(* Logix 5000 project; controller MV vendor 1 type 14 code 217 rev 31.11; software revision 31.00; part 42 of 53 *)
(* tags used below, declared in another part *)
   Always_Off : BOOL;
   Dummy : BOOL;
   MV20_TP_Capture_Volume_Timer : TIMER;
   MV_BM01_AV01_CIP : BOOL;
   MV_data_file_value_to_move : DINT;
   MV_Enable_MV20_NewPressureControl : BOOL;
   MV_from_data_file : DINT;
   MV_from_data_offset : DINT;
   MV_MV10_RTD1_AI : PlantItem;   // MV10_RTD1
   MV_MV11_RTD1_AI : PlantItem;   // MV11_RTD1
   MV_MV12_RTD1_AI : PlantItem;   // MV12_RTD1
   MV_MV13_RTD1_AI : PlantItem;   // MV13_RTD1
   MV_MV14_RTD1_AI : PlantItem;   // MV14_RTD1
   MV_MV15_RTD1_AI : PlantItem;   // MV15_RTD1
   MV_MV16_RTD1_AI : PlantItem;   // MV16_RTD1
   MV_MV17_RTD1_AI : PlantItem;   // MV17_RTD1
   MV_MV18_RTD1_AI : PlantItem;   // MV18_RTD1
   MV_MV19_RTD1_AI : PlantItem;   // MV19_RTD1
   MV_MV1_RTD1_AI : PlantItem;   // MV1_RTD1
   MV_MV20_CO2_ON_PreStorage : BOOL;
   MV_MV20_CO2_ON_Storage : BOOL;
   MV_MV20_Filling_PulseLevel : REAL;
   MV_MV20_LTX07_TrueLevel : REAL;
   MV_MV20_ProxiesOK : BOOL;
   MV_MV20_PTX01_AI : PlantItem;   // MV20_PTX01
   MV_MV20_RTD1_AI : PlantItem;   // MV20_RTD1
   MV_MV20_TP_Command : DINT;
   MV_MV20_TP_Dirty : BOOL;
   MV_MV20_TP_Emptying_Level_Setpoint : REAL;
   MV_MV20_TP_Idle : BOOL;
   MV_MV20_TP_KBDepressure : BOOL;
   MV_MV20_TP_KBFilling : BOOL;
   MV_MV20_TP_KBFilling_M : BOOL;
   MV_MV20_TP_KBPreEmptyPressure : BOOL;
   MV_MV20_TP_KBPrePressurise : BOOL;
   MV_MV20_TP_KBPurgeFromTop : BOOL;
   MV_MV20_TP_KBPurgeTimer : TIMER;
   MV_MV20_TP_KBStorage : BOOL;
   MV_MV20_TP_ONS : BOOL;
   MV_MV20_TP_Prompt : DINT;
   MV_MV20_TP_ReadyToFillKB : BOOL;
   MV_MV20_TP_ReadyToFillKB_M : BOOL;
   MV_MV20_TP_Running : BOOL;
   MV_MV20_TP_Setpoint : REAL;
   MV_MV20_TP_Status : DINT;   // 0 = Idle, 1 = Running, 2 = Held, 3 = Faulted
   MV_MV20_TP_Step : DINT;
   MV_MV20_TP_Steptime : DINT;
   MV_MV20_TP_UpperLimit : REAL;
   MV_MV20_Transfer_StartLevel : REAL;
   MV_MV21_RTD1_AI : PlantItem;   // MV21_RTD1
   MV_MV22_RTD1_AI : PlantItem;   // MV22_RTD1
   MV_MV23_RTD1_AI : PlantItem;   // MV23_RTD1
   MV_MV2_RTD1_AI : PlantItem;   // MV2_RTD1
   MV_MV30_RTD1_AI : PlantItem;   // MV30_RTD1
   MV_MV31_RTD1_AI : PlantItem;   // MV31_RTD1
   MV_MV32_RTD1_AI : PlantItem;   // MV32_RTD1
   MV_MV33_RTD1_AI : PlantItem;   // MV33_RTD1
   MV_MV34_RTD1_AI : PlantItem;   // MV34_RTD1
   MV_MV35_RTD1_AI : PlantItem;   // MV35_RTD1
   MV_MV36_TTX01_AI : PlantItem;   // MV36_TTX01
   MV_MV37_TTX01_AI : PlantItem;   // MV37_TTX01
   MV_MV38_TTX01_AI : PlantItem;   // MV38_TTX01
   MV_MV39_TTX01_AI : PlantItem;   // MV39_TTX01
   MV_MV3_RTD1_AI : PlantItem;   // MV3_RTD1
   MV_MV40_TTX01_AI : PlantItem;   // MV40_TTX01
   MV_MV41_TTX01_AI : PlantItem;   // MV41_TTX01
   MV_MV42_TTX01_AI : PlantItem;   // MV42_TTX01
   MV_MV43_TTX01_AI : PlantItem;   // MV43_TTX01
   MV_MV44_TTX01_AI : PlantItem;   // MV44_TTX01
   MV_MV45_TTX01_AI : PlantItem;   // MV45_TTX01
   MV_MV46_TTX01_AI : PlantItem;   // MV46_TTX01
   MV_MV47_TTX01_AI : PlantItem;   // MV47_TTX01
   MV_MV4_RTD1_AI : PlantItem;   // MV4_RTD1
   MV_MV5_RTD1_AI : PlantItem;   // MV5_RTD1
   MV_MV6_RTD1_AI : PlantItem;   // MV6_RTD1
   MV_MV7_RTD1_AI : PlantItem;   // MV7_RTD1
   MV_MV8_RTD1_AI : PlantItem;   // MV8_RTD1
   MV_MV9_RTD1_AI : PlantItem;   // MV9_RTD1
   MV_N106 : INT[255];   // ROUSE_BUFF Rouser control vesse l data buffer
   MV_N110 : INT[255];   // MV DATA 0 CURRENT FV DATA
   MV_N111 : INT[50];   // MV 1, CURRENT FV DATA
   MV_N112 : INT[50];   // MV 2, CURRENT FV DATA
   MV_N113 : INT[50];   // MV 3, CURRENT FV DATA
   MV_N114 : INT[50];   // MV 4, CURRENT FV DATA
   MV_N115 : INT[50];   // MV 5, CURRENT FV DATA
   MV_N116 : INT[50];   // MV 6, CURRENT FV DATA
   MV_N117 : INT[50];   // MV 7, CURRENT FV DATA
   MV_N118 : INT[50];   // MV 8, CURRENT FV DATA
   MV_N119 : INT[50];   // MV 9, CURRENT FV DATA
   MV_N120 : INT[50];   // MV 10, CURRENT FV DATA
   MV_N121 : INT[50];   // MV 11, CURRENT FV DATA
   MV_N122 : INT[50];   // MV 12, CURRENT FV DATA
   MV_N123 : INT[50];   // MV 13, CURRENT FV DATA
   MV_N124 : INT[50];   // MV 14, CURRENT FV DATA
   MV_N125 : INT[50];   // MV 15, CURRENT FV DATA
   MV_N126 : INT[50];   // MV 16, CURRENT FV DATA
   MV_N127 : INT[50];   // MV 17, CURRENT FV DATA
   MV_N128 : INT[50];   // MV 18, CURRENT FV DATA
   MV_N129 : INT[50];   // MV 19, CURRENT FV DATA
   MV_N130 : INT[50];   // MV 30, CURRENT FV DATA
   MV_N131 : INT[50];   // MV 31, CURRENT FV DATA
   MV_N132 : INT[50];   // MV 32, CURRENT FV DATA
   MV_N133 : INT[50];   // MV 33, CURRENT FV DATA
   MV_N134 : INT[50];   // MV 34, CURRENT FV DATA
   MV_N135 : INT[50];   // MV 35, CURRENT FV DATA
   MV_N136 : INT[50];   // MV 20, CURRENT FV DATA
   MV_N137 : INT[50];   // MV 21, CURRENT FV DATA
   MV_N138 : INT[50];   // MV 22, CURRENT FV DATA
   MV_N139 : INT[50];   // MV 23, CURRENT FV DATA
   MV_N140 : INT[50];   // MV 36, CURRENT FV DATA
   MV_N141 : INT[50];   // MV 37, CURRENT FV DATA
   MV_N142 : INT[50];   // MV 38, CURRENT FV DATA
   MV_N143 : INT[50];   // MV 39, CURRENT FV DATA
   MV_N144 : INT[50];   // MV 40, CURRENT FV DATA
   MV_N145 : INT[50];   // MV 41, CURRENT FV DATA
   MV_N146 : INT[50];   // MV 42, CURRENT FV DATA
   MV_N147 : INT[50];   // MV 43, CURRENT FV DATA
   MV_N148 : INT[50];   // MV 44, CURRENT FV DATA
   MV_N149 : INT[50];   // MV 45, CURRENT FV DATA
   MV_N150 : INT[50];   // MV 36, CURRENT FV DATA
   MV_N151 : INT[50];   // MV 47, CURRENT FV DATA
   MV_TP_CaskPrefillPressure : REAL;
   MV_TP_Emptying_Volume_Setpoint : REAL;
   MV_TP_KBEmptyingPressure : REAL;
   MV_TP_KBFillingPressure : REAL;
   MV_TP_KBPrefillPressure : REAL;
   MV_TP_KBStoragePressure : REAL;
   MV_TP_KBStoragePressureLevel : REAL;
   MV_TP_NoCIPDelay : DINT;
(* MV_Common, continued *)

ROUTINE MV_Get_FV_Datafile_Value   (* ladder *)
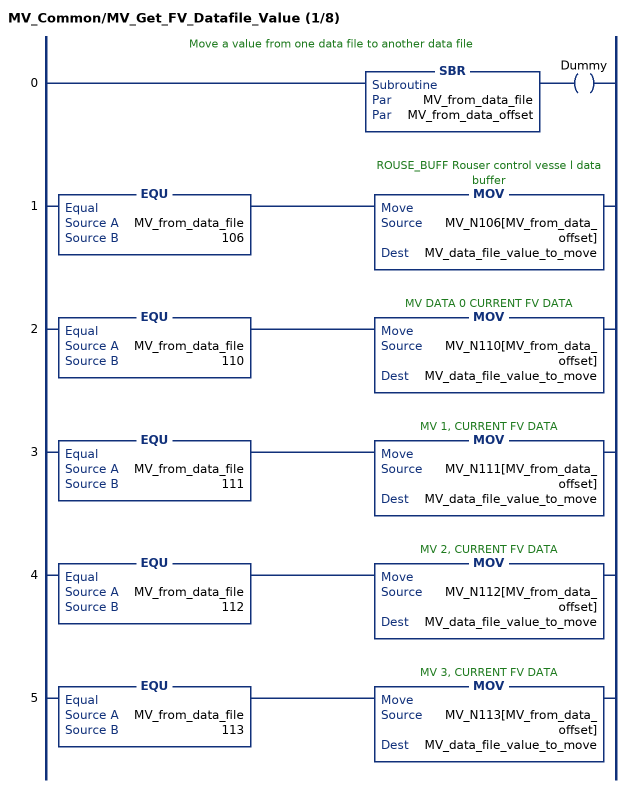
   // Move a value from one data file to another data file
   0: SBR(MV_from_data_file,MV_from_data_offset)OTE(Dummy);
   1: EQU(MV_from_data_file,106)MOV(MV_N106[MV_from_data_offset],MV_data_file_value_to_move);
   2: EQU(MV_from_data_file,110)MOV(MV_N110[MV_from_data_offset],MV_data_file_value_to_move);
   3: EQU(MV_from_data_file,111)MOV(MV_N111[MV_from_data_offset],MV_data_file_value_to_move);
   4: EQU(MV_from_data_file,112)MOV(MV_N112[MV_from_data_offset],MV_data_file_value_to_move);
   5: EQU(MV_from_data_file,113)MOV(MV_N113[MV_from_data_offset],MV_data_file_value_to_move);
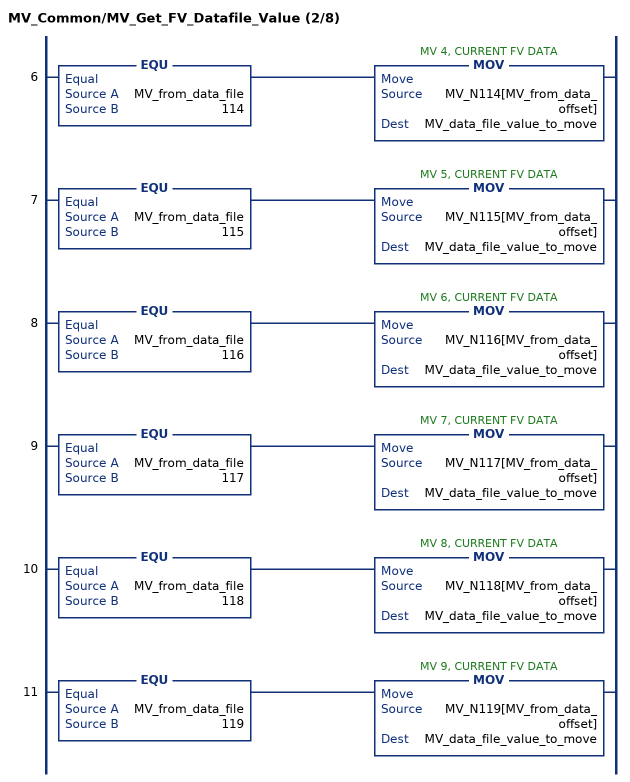
   6: EQU(MV_from_data_file,114)MOV(MV_N114[MV_from_data_offset],MV_data_file_value_to_move);
   7: EQU(MV_from_data_file,115)MOV(MV_N115[MV_from_data_offset],MV_data_file_value_to_move);
   8: EQU(MV_from_data_file,116)MOV(MV_N116[MV_from_data_offset],MV_data_file_value_to_move);
   9: EQU(MV_from_data_file,117)MOV(MV_N117[MV_from_data_offset],MV_data_file_value_to_move);
   10: EQU(MV_from_data_file,118)MOV(MV_N118[MV_from_data_offset],MV_data_file_value_to_move);
   11: EQU(MV_from_data_file,119)MOV(MV_N119[MV_from_data_offset],MV_data_file_value_to_move);
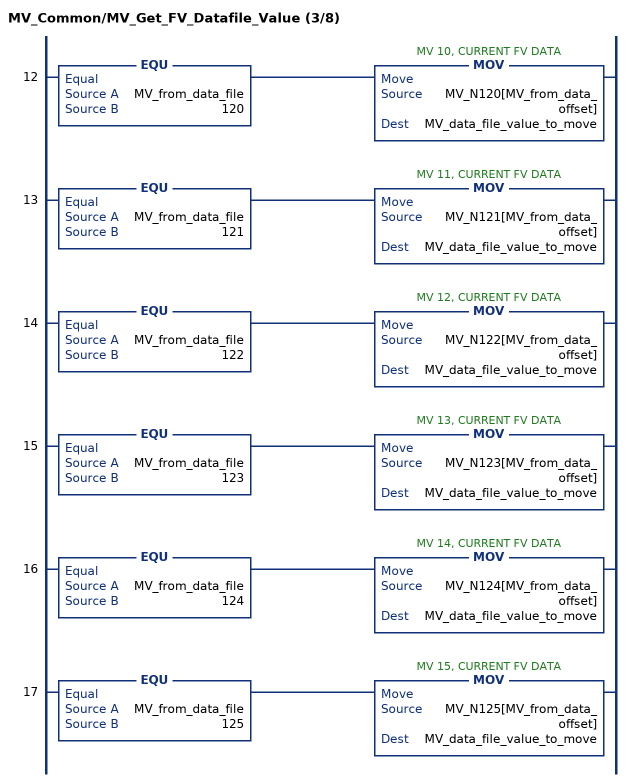
   12: EQU(MV_from_data_file,120)MOV(MV_N120[MV_from_data_offset],MV_data_file_value_to_move);
   13: EQU(MV_from_data_file,121)MOV(MV_N121[MV_from_data_offset],MV_data_file_value_to_move);
   14: EQU(MV_from_data_file,122)MOV(MV_N122[MV_from_data_offset],MV_data_file_value_to_move);
   15: EQU(MV_from_data_file,123)MOV(MV_N123[MV_from_data_offset],MV_data_file_value_to_move);
   16: EQU(MV_from_data_file,124)MOV(MV_N124[MV_from_data_offset],MV_data_file_value_to_move);
   17: EQU(MV_from_data_file,125)MOV(MV_N125[MV_from_data_offset],MV_data_file_value_to_move);
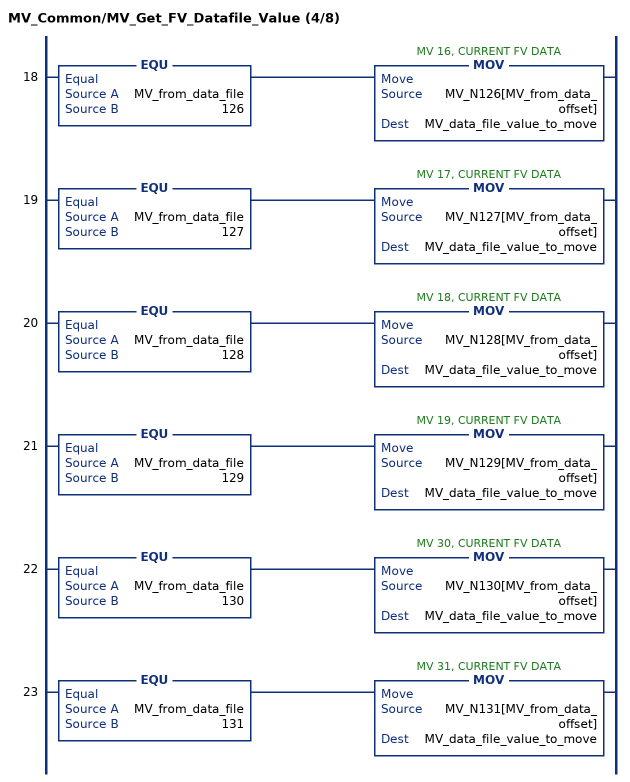
   18: EQU(MV_from_data_file,126)MOV(MV_N126[MV_from_data_offset],MV_data_file_value_to_move);
   19: EQU(MV_from_data_file,127)MOV(MV_N127[MV_from_data_offset],MV_data_file_value_to_move);
   20: EQU(MV_from_data_file,128)MOV(MV_N128[MV_from_data_offset],MV_data_file_value_to_move);
   21: EQU(MV_from_data_file,129)MOV(MV_N129[MV_from_data_offset],MV_data_file_value_to_move);
   22: EQU(MV_from_data_file,130)MOV(MV_N130[MV_from_data_offset],MV_data_file_value_to_move);
   23: EQU(MV_from_data_file,131)MOV(MV_N131[MV_from_data_offset],MV_data_file_value_to_move);
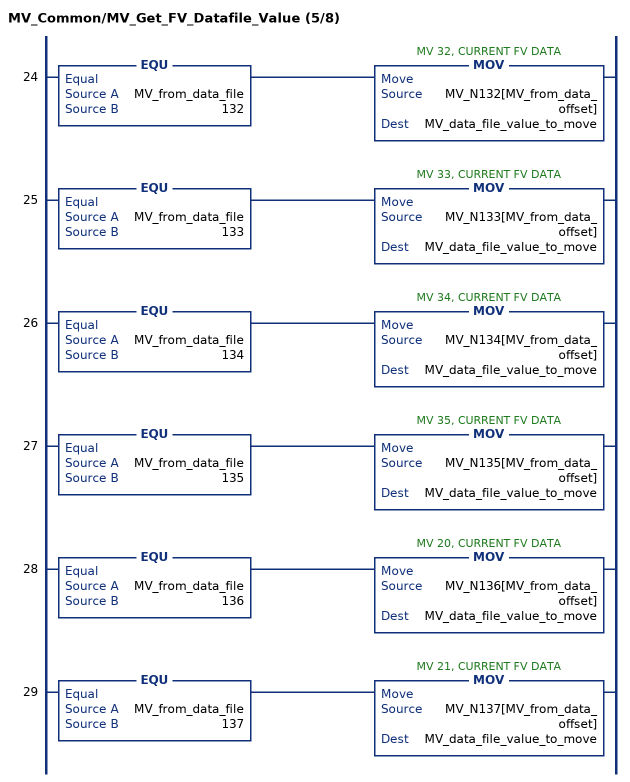
   24: EQU(MV_from_data_file,132)MOV(MV_N132[MV_from_data_offset],MV_data_file_value_to_move);
   25: EQU(MV_from_data_file,133)MOV(MV_N133[MV_from_data_offset],MV_data_file_value_to_move);
   26: EQU(MV_from_data_file,134)MOV(MV_N134[MV_from_data_offset],MV_data_file_value_to_move);
   27: EQU(MV_from_data_file,135)MOV(MV_N135[MV_from_data_offset],MV_data_file_value_to_move);
   28: EQU(MV_from_data_file,136)MOV(MV_N136[MV_from_data_offset],MV_data_file_value_to_move);
   29: EQU(MV_from_data_file,137)MOV(MV_N137[MV_from_data_offset],MV_data_file_value_to_move);
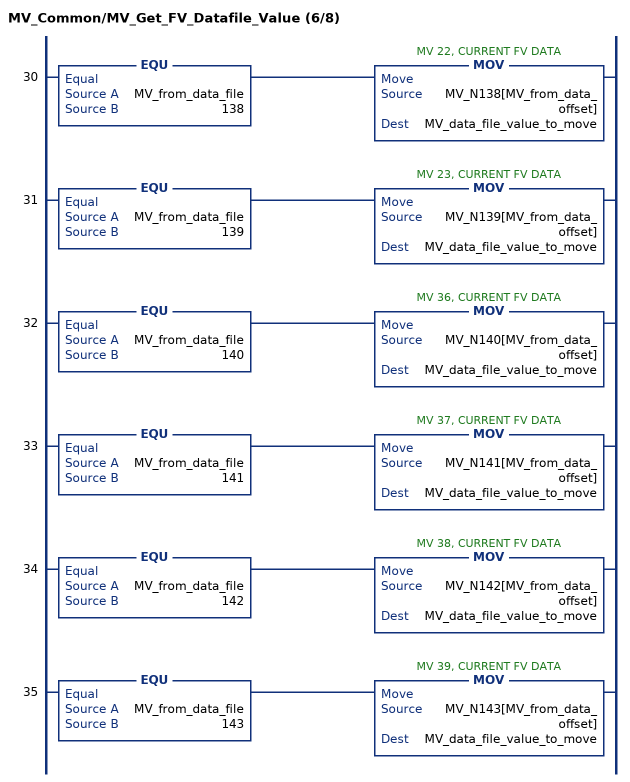
   30: EQU(MV_from_data_file,138)MOV(MV_N138[MV_from_data_offset],MV_data_file_value_to_move);
   31: EQU(MV_from_data_file,139)MOV(MV_N139[MV_from_data_offset],MV_data_file_value_to_move);
   32: EQU(MV_from_data_file,140)MOV(MV_N140[MV_from_data_offset],MV_data_file_value_to_move);
   33: EQU(MV_from_data_file,141)MOV(MV_N141[MV_from_data_offset],MV_data_file_value_to_move);
   34: EQU(MV_from_data_file,142)MOV(MV_N142[MV_from_data_offset],MV_data_file_value_to_move);
   35: EQU(MV_from_data_file,143)MOV(MV_N143[MV_from_data_offset],MV_data_file_value_to_move);
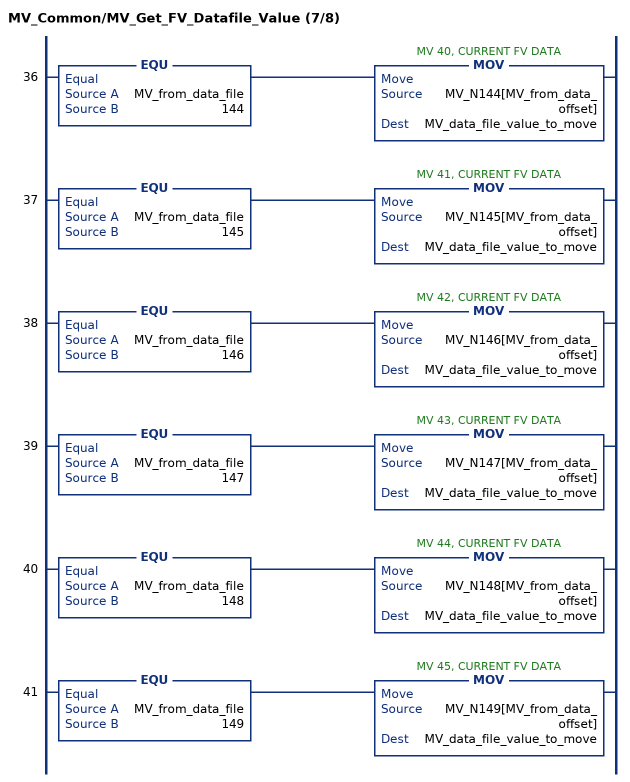
   36: EQU(MV_from_data_file,144)MOV(MV_N144[MV_from_data_offset],MV_data_file_value_to_move);
   37: EQU(MV_from_data_file,145)MOV(MV_N145[MV_from_data_offset],MV_data_file_value_to_move);
   38: EQU(MV_from_data_file,146)MOV(MV_N146[MV_from_data_offset],MV_data_file_value_to_move);
   39: EQU(MV_from_data_file,147)MOV(MV_N147[MV_from_data_offset],MV_data_file_value_to_move);
   40: EQU(MV_from_data_file,148)MOV(MV_N148[MV_from_data_offset],MV_data_file_value_to_move);
   41: EQU(MV_from_data_file,149)MOV(MV_N149[MV_from_data_offset],MV_data_file_value_to_move);
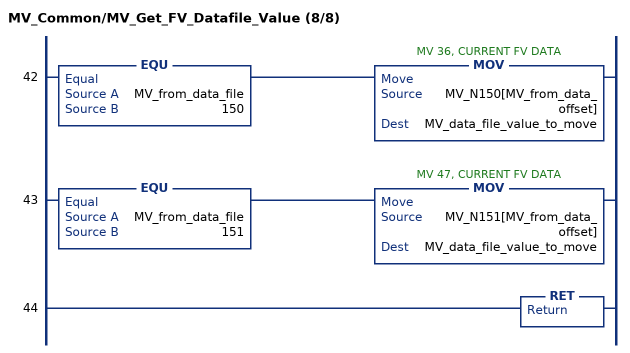
   42: EQU(MV_from_data_file,150)MOV(MV_N150[MV_from_data_offset],MV_data_file_value_to_move);
   43: EQU(MV_from_data_file,151)MOV(MV_N151[MV_from_data_offset],MV_data_file_value_to_move);
   44: RET();
END_ROUTINE

ROUTINE MV_Move_Temps_To_DataFiles   (* ladder *)
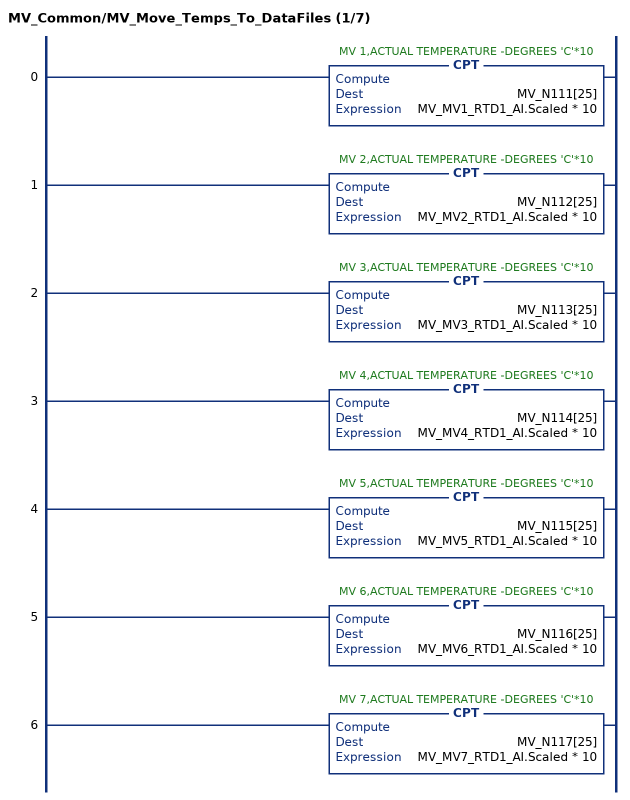
   0: CPT(MV_N111[25],MV_MV1_RTD1_AI.Scaled * 10);
   1: CPT(MV_N112[25],MV_MV2_RTD1_AI.Scaled * 10);
   2: CPT(MV_N113[25],MV_MV3_RTD1_AI.Scaled * 10);
   3: CPT(MV_N114[25],MV_MV4_RTD1_AI.Scaled * 10);
   4: CPT(MV_N115[25],MV_MV5_RTD1_AI.Scaled * 10);
   5: CPT(MV_N116[25],MV_MV6_RTD1_AI.Scaled * 10);
   6: CPT(MV_N117[25],MV_MV7_RTD1_AI.Scaled * 10);
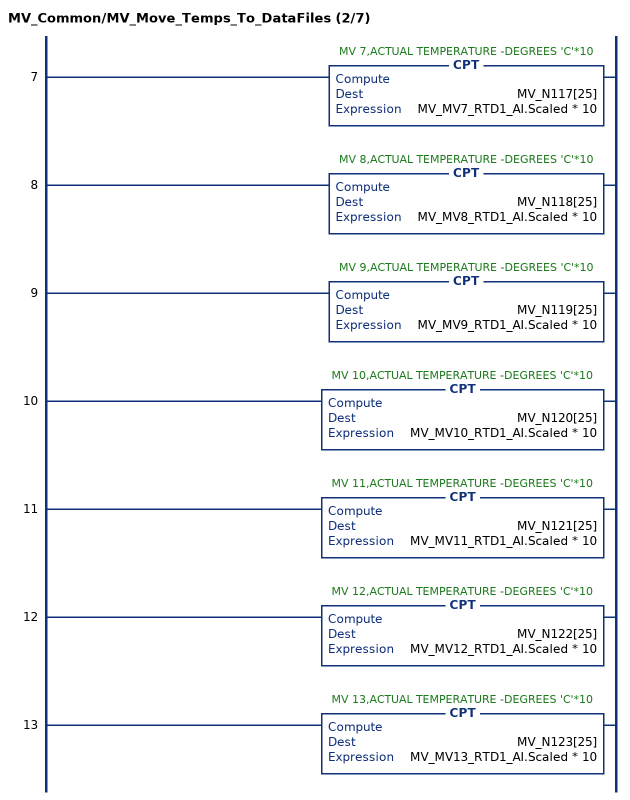
   7: CPT(MV_N117[25],MV_MV7_RTD1_AI.Scaled * 10);
   8: CPT(MV_N118[25],MV_MV8_RTD1_AI.Scaled * 10);
   9: CPT(MV_N119[25],MV_MV9_RTD1_AI.Scaled * 10);
   10: CPT(MV_N120[25],MV_MV10_RTD1_AI.Scaled * 10);
   11: CPT(MV_N121[25],MV_MV11_RTD1_AI.Scaled * 10);
   12: CPT(MV_N122[25],MV_MV12_RTD1_AI.Scaled * 10);
   13: CPT(MV_N123[25],MV_MV13_RTD1_AI.Scaled * 10);
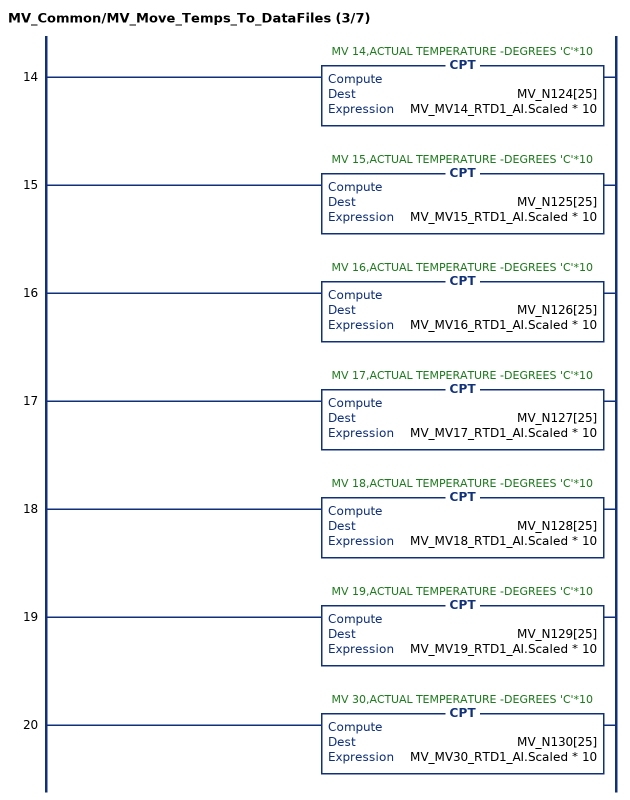
   14: CPT(MV_N124[25],MV_MV14_RTD1_AI.Scaled * 10);
   15: CPT(MV_N125[25],MV_MV15_RTD1_AI.Scaled * 10);
   16: CPT(MV_N126[25],MV_MV16_RTD1_AI.Scaled * 10);
   17: CPT(MV_N127[25],MV_MV17_RTD1_AI.Scaled * 10);
   18: CPT(MV_N128[25],MV_MV18_RTD1_AI.Scaled * 10);
   19: CPT(MV_N129[25],MV_MV19_RTD1_AI.Scaled * 10);
   20: CPT(MV_N130[25],MV_MV30_RTD1_AI.Scaled * 10);
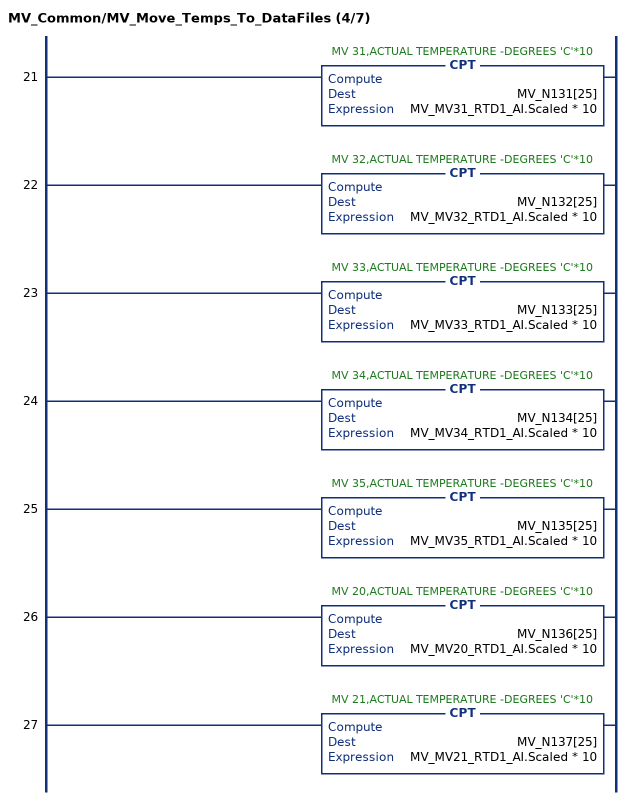
   21: CPT(MV_N131[25],MV_MV31_RTD1_AI.Scaled * 10);
   22: CPT(MV_N132[25],MV_MV32_RTD1_AI.Scaled * 10);
   23: CPT(MV_N133[25],MV_MV33_RTD1_AI.Scaled * 10);
   24: CPT(MV_N134[25],MV_MV34_RTD1_AI.Scaled * 10);
   25: CPT(MV_N135[25],MV_MV35_RTD1_AI.Scaled * 10);
   26: CPT(MV_N136[25],MV_MV20_RTD1_AI.Scaled * 10);
   27: CPT(MV_N137[25],MV_MV21_RTD1_AI.Scaled * 10);
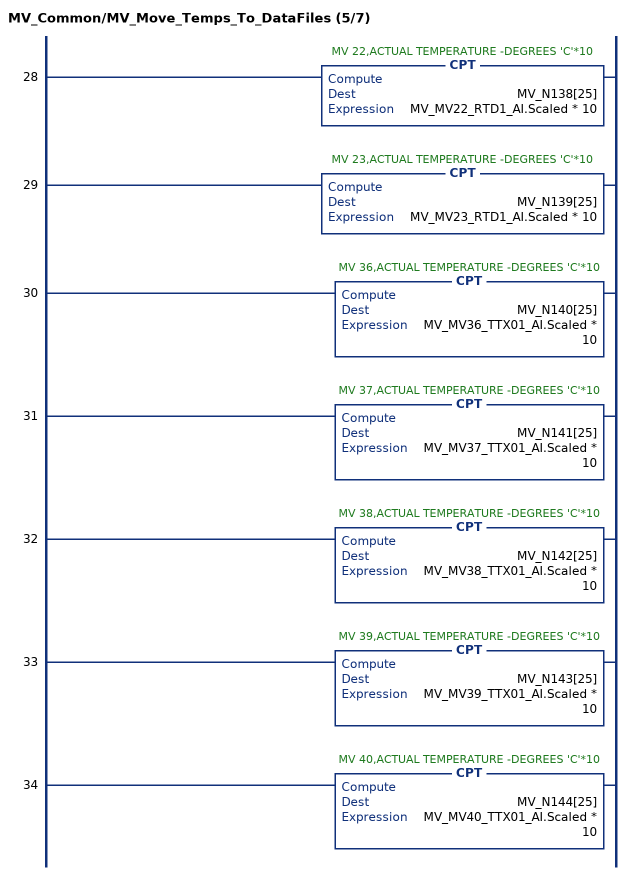
   28: CPT(MV_N138[25],MV_MV22_RTD1_AI.Scaled * 10);
   29: CPT(MV_N139[25],MV_MV23_RTD1_AI.Scaled * 10);
   30: CPT(MV_N140[25],MV_MV36_TTX01_AI.Scaled * 10);
   31: CPT(MV_N141[25],MV_MV37_TTX01_AI.Scaled * 10);
   32: CPT(MV_N142[25],MV_MV38_TTX01_AI.Scaled * 10);
   33: CPT(MV_N143[25],MV_MV39_TTX01_AI.Scaled * 10);
   34: CPT(MV_N144[25],MV_MV40_TTX01_AI.Scaled * 10);
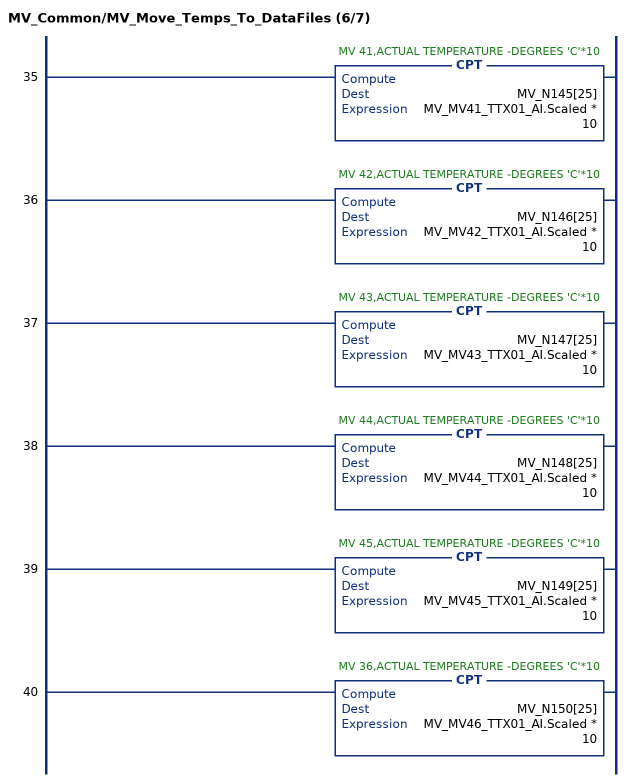
   35: CPT(MV_N145[25],MV_MV41_TTX01_AI.Scaled * 10);
   36: CPT(MV_N146[25],MV_MV42_TTX01_AI.Scaled * 10);
   37: CPT(MV_N147[25],MV_MV43_TTX01_AI.Scaled * 10);
   38: CPT(MV_N148[25],MV_MV44_TTX01_AI.Scaled * 10);
   39: CPT(MV_N149[25],MV_MV45_TTX01_AI.Scaled * 10);
   40: CPT(MV_N150[25],MV_MV46_TTX01_AI.Scaled * 10);
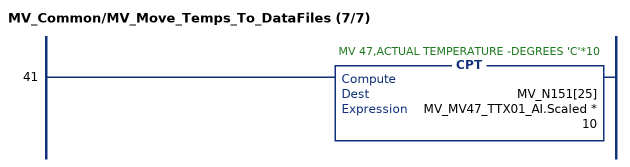
   41: CPT(MV_N151[25],MV_MV47_TTX01_AI.Scaled * 10);
END_ROUTINE

ROUTINE MV_MV20_TP   (* ladder *)
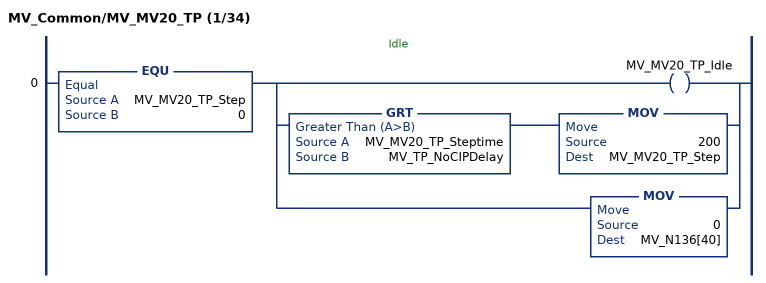
   // Idle
   0: EQU(MV_MV20_TP_Step,0)[OTE(MV_MV20_TP_Idle) ,GRT(MV_MV20_TP_Steptime,MV_TP_NoCIPDelay) MOV(200,MV_MV20_TP_Step) ,MOV(0,MV_N136[40]) ];
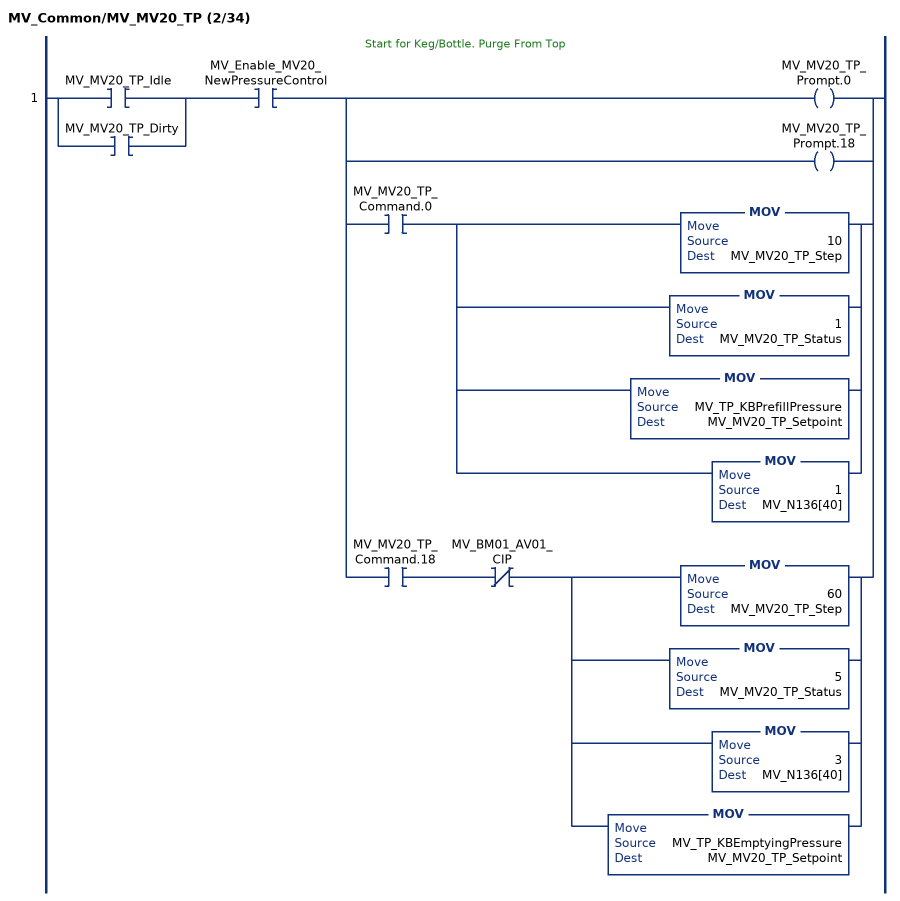
   // Start for Keg/Bottle. Purge From Top
   1: [XIC(MV_MV20_TP_Idle) ,XIC(MV_MV20_TP_Dirty) ]XIC(MV_Enable_MV20_NewPressureControl)[OTE(MV_MV20_TP_Prompt.0) ,OTE(MV_MV20_TP_Prompt.18) ,XIC(MV_MV20_TP_Command.0) [MOV(10,MV_MV20_TP_Step) ,MOV(1,MV_MV20_TP_Status) ,MOV(MV_TP_KBPrefillPressure,MV_MV20_TP_Setpoint) ,MOV(1,MV_N136[40]) ] ,XIC(MV_MV20_TP_Command.18) XIO(MV_BM01_AV01_CIP) [MOV(60,MV_MV20_TP_Step) ,MOV(5,MV_MV20_TP_Status) ,MOV(3,MV_N136[40]) ,MOV(MV_TP_KBEmptyingPressure,MV_MV20_TP_Setpoint) ] ];
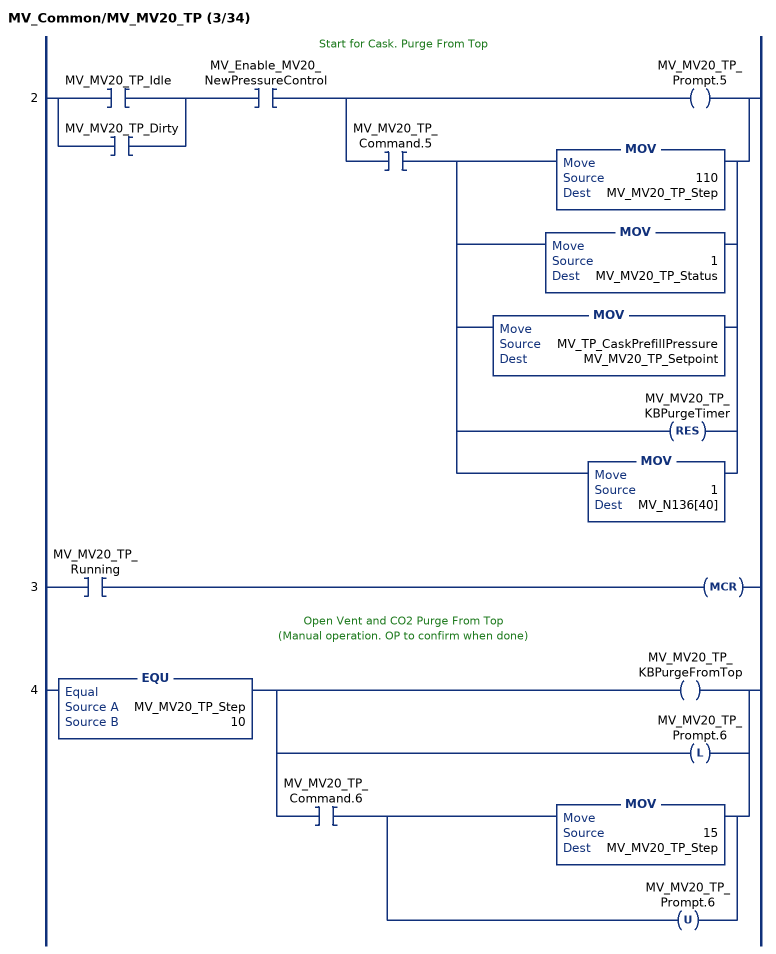
   // Start for Cask. Purge From Top
   2: [XIC(MV_MV20_TP_Idle) ,XIC(MV_MV20_TP_Dirty) ]XIC(MV_Enable_MV20_NewPressureControl)[OTE(MV_MV20_TP_Prompt.5) ,XIC(MV_MV20_TP_Command.5) [MOV(110,MV_MV20_TP_Step) ,MOV(1,MV_MV20_TP_Status) ,MOV(MV_TP_CaskPrefillPressure,MV_MV20_TP_Setpoint) ,RES(MV_MV20_TP_KBPurgeTimer) ,MOV(1,MV_N136[40]) ] ];
   3: XIC(MV_MV20_TP_Running)MCR();
   // Open Vent and CO2 Purge From Top
   // (Manual operation. OP to confirm when done)
   4: EQU(MV_MV20_TP_Step,10)[OTE(MV_MV20_TP_KBPurgeFromTop) ,OTL(MV_MV20_TP_Prompt.6) ,XIC(MV_MV20_TP_Command.6) [MOV(15,MV_MV20_TP_Step) ,OTU(MV_MV20_TP_Prompt.6) ] ];
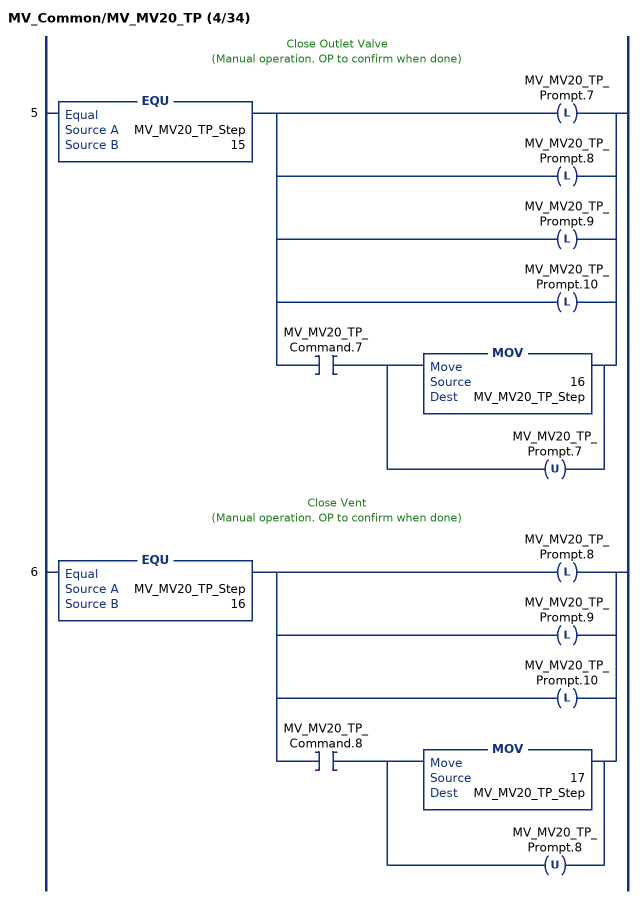
   // Close Outlet Valve
   // (Manual operation. OP to confirm when done)
   5: EQU(MV_MV20_TP_Step,15)[OTL(MV_MV20_TP_Prompt.7) ,OTL(MV_MV20_TP_Prompt.8) ,OTL(MV_MV20_TP_Prompt.9) ,OTL(MV_MV20_TP_Prompt.10) ,XIC(MV_MV20_TP_Command.7) [MOV(16,MV_MV20_TP_Step) ,OTU(MV_MV20_TP_Prompt.7) ] ];
   // Close Vent
   // (Manual operation. OP to confirm when done)
   6: EQU(MV_MV20_TP_Step,16)[OTL(MV_MV20_TP_Prompt.8) ,OTL(MV_MV20_TP_Prompt.9) ,OTL(MV_MV20_TP_Prompt.10) ,XIC(MV_MV20_TP_Command.8) [MOV(17,MV_MV20_TP_Step) ,OTU(MV_MV20_TP_Prompt.8) ] ];
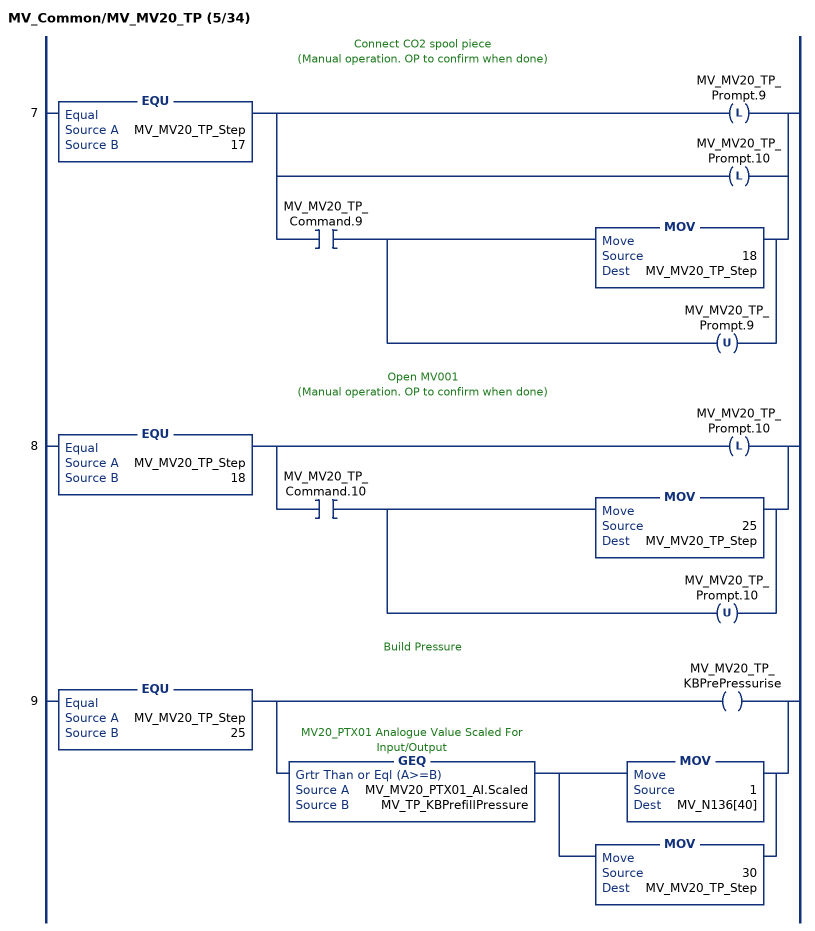
   // Connect CO2 spool piece
   // (Manual operation. OP to confirm when done)
   7: EQU(MV_MV20_TP_Step,17)[OTL(MV_MV20_TP_Prompt.9) ,OTL(MV_MV20_TP_Prompt.10) ,XIC(MV_MV20_TP_Command.9) [MOV(18,MV_MV20_TP_Step) ,OTU(MV_MV20_TP_Prompt.9) ] ];
   // Open MV001
   // (Manual operation. OP to confirm when done)
   8: EQU(MV_MV20_TP_Step,18)[OTL(MV_MV20_TP_Prompt.10) ,XIC(MV_MV20_TP_Command.10) [MOV(25,MV_MV20_TP_Step) ,OTU(MV_MV20_TP_Prompt.10) ] ];
   // Build Pressure
   9: EQU(MV_MV20_TP_Step,25)[OTE(MV_MV20_TP_KBPrePressurise) ,GEQ(MV_MV20_PTX01_AI.Scaled,MV_TP_KBPrefillPressure) [MOV(1,MV_N136[40]) ,MOV(30,MV_MV20_TP_Step) ] ];
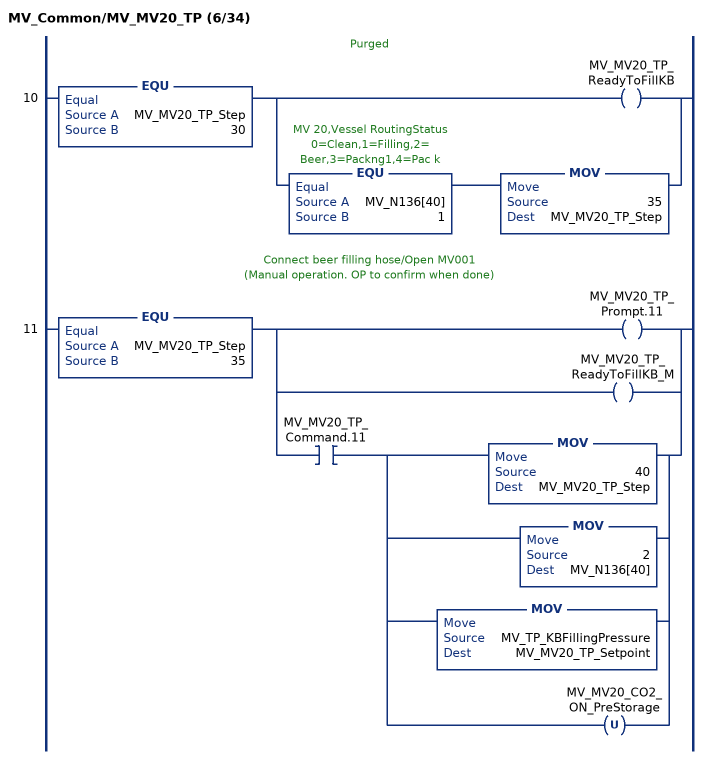
   // Purged
   10: EQU(MV_MV20_TP_Step,30)[OTE(MV_MV20_TP_ReadyToFillKB) ,EQU(MV_N136[40],1) MOV(35,MV_MV20_TP_Step) ];
   // Connect beer filling hose/Open MV001
   // (Manual operation. OP to confirm when done)
   11: EQU(MV_MV20_TP_Step,35)[OTE(MV_MV20_TP_Prompt.11) ,OTE(MV_MV20_TP_ReadyToFillKB_M) ,XIC(MV_MV20_TP_Command.11) [MOV(40,MV_MV20_TP_Step) ,MOV(2,MV_N136[40]) ,MOV(MV_TP_KBFillingPressure,MV_MV20_TP_Setpoint) ,OTU(MV_MV20_CO2_ON_PreStorage) ] ];
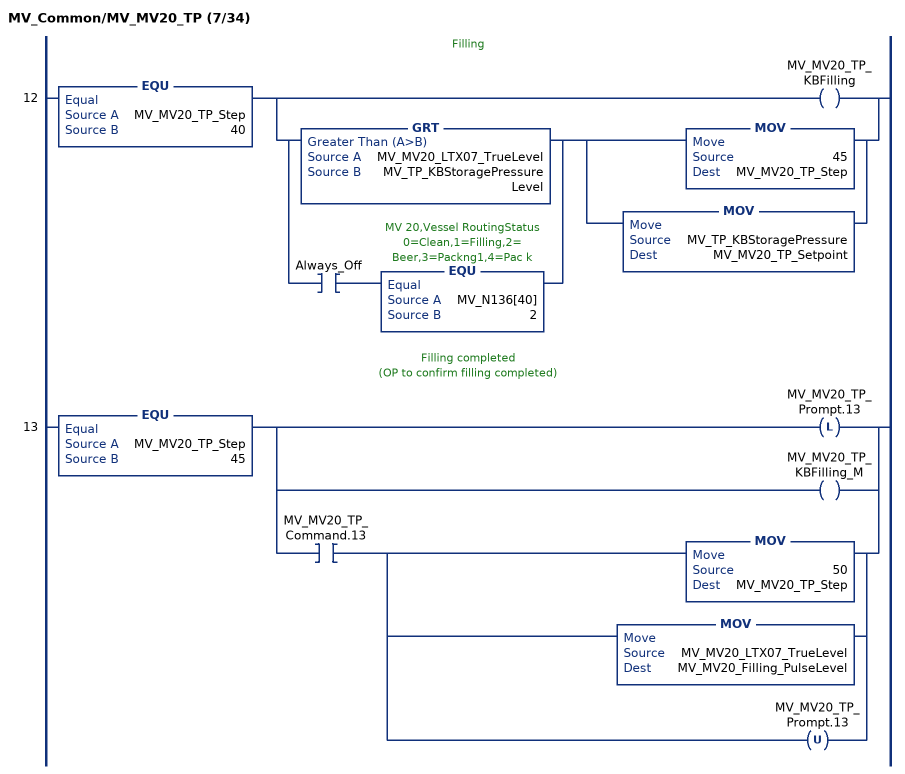
   // Filling
   12: EQU(MV_MV20_TP_Step,40)[OTE(MV_MV20_TP_KBFilling) ,[GRT(MV_MV20_LTX07_TrueLevel,MV_TP_KBStoragePressureLevel) ,XIC(Always_Off) EQU(MV_N136[40],2) ] [MOV(45,MV_MV20_TP_Step) ,MOV(MV_TP_KBStoragePressure,MV_MV20_TP_Setpoint) ] ];
   // Filling completed
   // (OP to confirm filling completed)
   13: EQU(MV_MV20_TP_Step,45)[OTL(MV_MV20_TP_Prompt.13) ,OTE(MV_MV20_TP_KBFilling_M) ,XIC(MV_MV20_TP_Command.13) [MOV(50,MV_MV20_TP_Step) ,MOV(MV_MV20_LTX07_TrueLevel,MV_MV20_Filling_PulseLevel) ,OTU(MV_MV20_TP_Prompt.13) ] ];
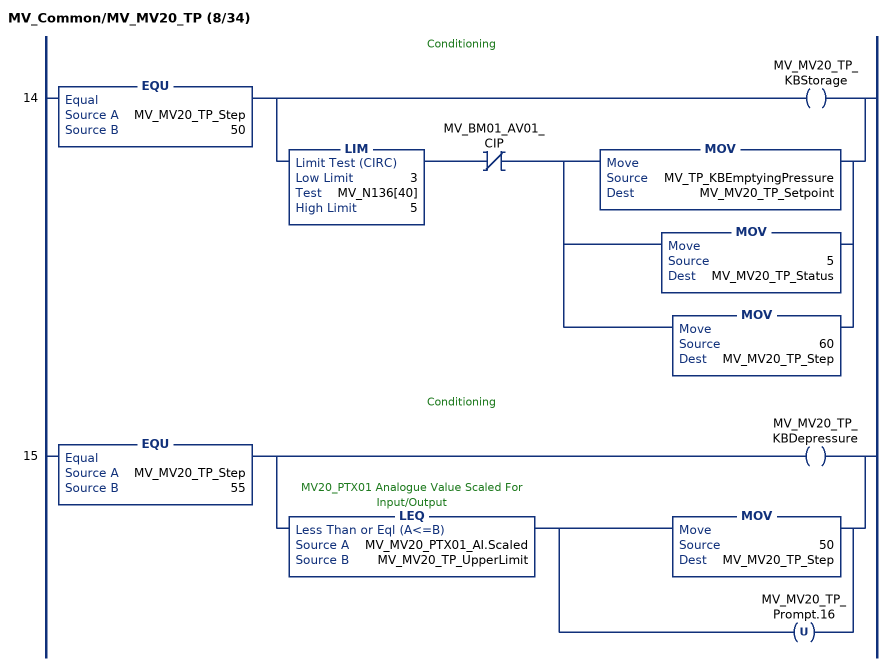
   // Conditioning
   14: EQU(MV_MV20_TP_Step,50)[OTE(MV_MV20_TP_KBStorage) ,LIM(3,MV_N136[40],5) XIO(MV_BM01_AV01_CIP) [MOV(MV_TP_KBEmptyingPressure,MV_MV20_TP_Setpoint) ,MOV(5,MV_MV20_TP_Status) ,MOV(60,MV_MV20_TP_Step) ] ];
   // Conditioning
   15: EQU(MV_MV20_TP_Step,55)[OTE(MV_MV20_TP_KBDepressure) ,LEQ(MV_MV20_PTX01_AI.Scaled,MV_MV20_TP_UpperLimit) [MOV(50,MV_MV20_TP_Step) ,OTU(MV_MV20_TP_Prompt.16) ] ];
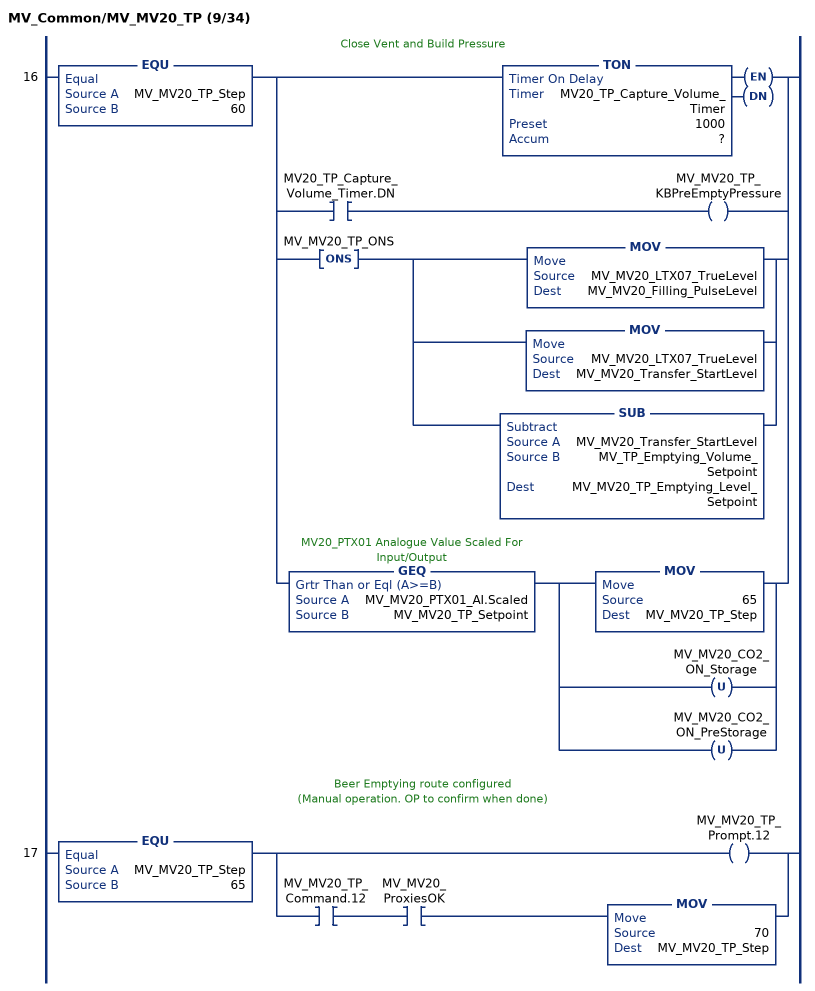
   // Close Vent and Build Pressure
   16: EQU(MV_MV20_TP_Step,60)[TON(MV20_TP_Capture_Volume_Timer,?,?) ,XIC(MV20_TP_Capture_Volume_Timer.DN) OTE(MV_MV20_TP_KBPreEmptyPressure) ,ONS(MV_MV20_TP_ONS) [MOV(MV_MV20_LTX07_TrueLevel,MV_MV20_Filling_PulseLevel) ,MOV(MV_MV20_LTX07_TrueLevel,MV_MV20_Transfer_StartLevel) ,SUB(MV_MV20_Transfer_StartLevel,MV_TP_Emptying_Volume_Setpoint,MV_MV20_TP_Emptying_Level_Setpoint) ] ,GEQ(MV_MV20_PTX01_AI.Scaled,MV_MV20_TP_Setpoint) [MOV(65,MV_MV20_TP_Step) ,OTU(MV_MV20_CO2_ON_Storage) ,OTU(MV_MV20_CO2_ON_PreStorage) ] ];
   // Beer Emptying route configured
   // (Manual operation. OP to confirm when done)
   17: EQU(MV_MV20_TP_Step,65)[OTE(MV_MV20_TP_Prompt.12) ,XIC(MV_MV20_TP_Command.12) XIC(MV_MV20_ProxiesOK) MOV(70,MV_MV20_TP_Step) ];
